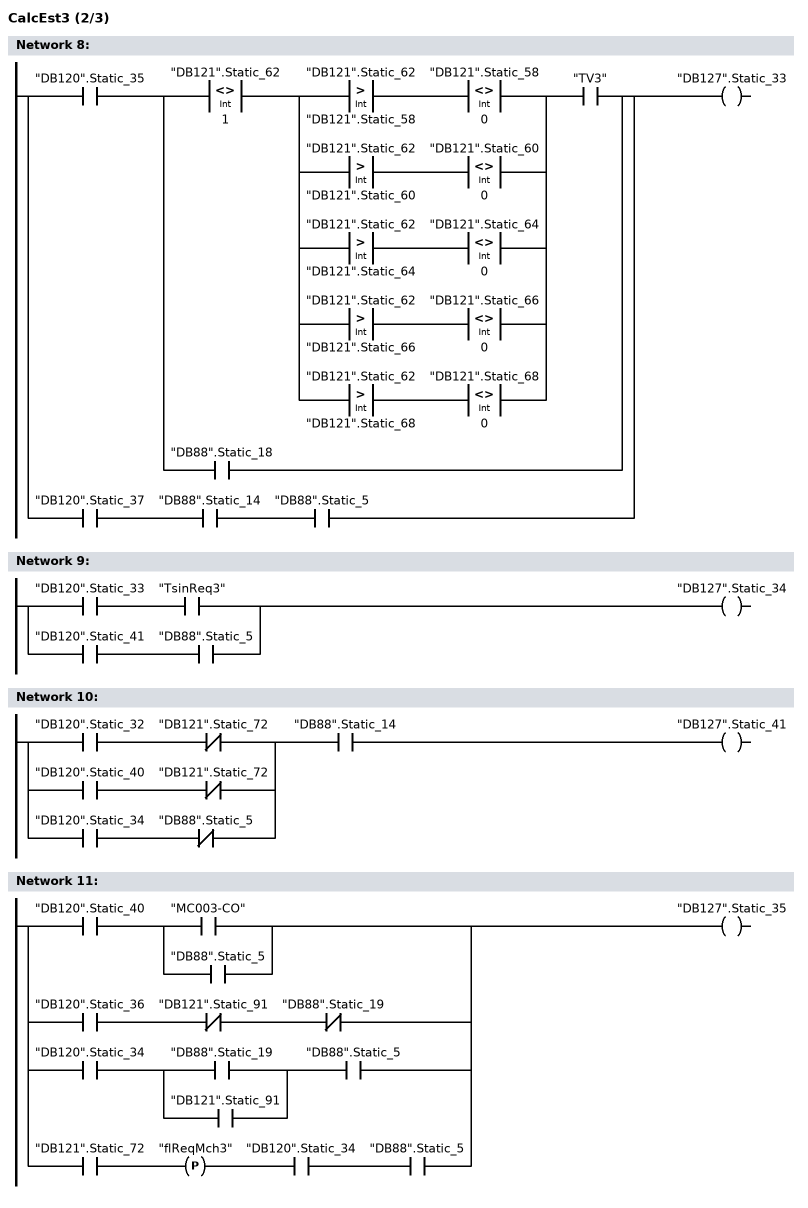
   "DB127".Static_33 := ("DB120".Static_35 AND ((("DB121".Static_62 <> 1) AND ((("DB121".Static_62 > "DB121".Static_58) AND ("DB121".Static_58 <> 0)) OR (("DB121".Static_62 > "DB121".Static_60) AND ("DB121".Static_60 <> 0)) OR (("DB121".Static_62 > "DB121".Static_64) AND ("DB121".Static_64 <> 0)) OR (("DB121".Static_62 > "DB121".Static_66) AND ("DB121".Static_66 <> 0)) OR (("DB121".Static_62 > "DB121".Static_68) AND ("DB121".Static_68 <> 0))) AND "TV3") OR "DB88".Static_18)) OR ("DB120".Static_37 AND "DB88".Static_14 AND "DB88".Static_5);
END_REGION

REGION Network 9
   RUNG wire#powerrail
      Contact( "DB120".Static_33 )
      Contact( "TsinReq3" )
      wire#w1
      Coil( "DB127".Static_34 )
   END_RUNG
   RUNG wire#powerrail
      Contact( "DB120".Static_41 )
      Contact( "DB88".Static_5 )
   END_RUNG wire#w1
   // the same network as SCL:
   "DB127".Static_34 := ("DB120".Static_33 AND "TsinReq3") OR ("DB120".Static_41 AND "DB88".Static_5);
END_REGION

REGION Network 10
   RUNG wire#powerrail
      Contact( "DB120".Static_32 )
      I_Contact( "DB121".Static_72 )
      wire#w1
      Contact( "DB88".Static_14 )
      Coil( "DB127".Static_41 )
   END_RUNG
   RUNG wire#powerrail
      Contact( "DB120".Static_40 )
      I_Contact( "DB121".Static_72 )
   END_RUNG wire#w1
   RUNG wire#powerrail
      Contact( "DB120".Static_34 )
      I_Contact( "DB88".Static_5 )
   END_RUNG wire#w1
   // the same network as SCL:
   "DB127".Static_41 := (("DB120".Static_32 AND NOT "DB121".Static_72) OR ("DB120".Static_40 AND NOT "DB121".Static_72) OR ("DB120".Static_34 AND NOT "DB88".Static_5)) AND "DB88".Static_14;
END_REGION

REGION Network 11
   #_w1 := "DB121".Static_72 AND NOT "flReqMch3";   // rising edge
   "flReqMch3" := "DB121".Static_72;
   "DB127".Static_35 := ("DB120".Static_40 AND ("MC003-CO" OR "DB88".Static_5)) OR ("DB120".Static_36 AND NOT "DB121".Static_91 AND NOT "DB88".Static_19) OR ("DB120".Static_34 AND ("DB88".Static_19 OR "DB121".Static_91) AND "DB88".Static_5) OR (#_w1 AND "DB120".Static_34 AND "DB88".Static_5);
END_REGION

REGION Network 12
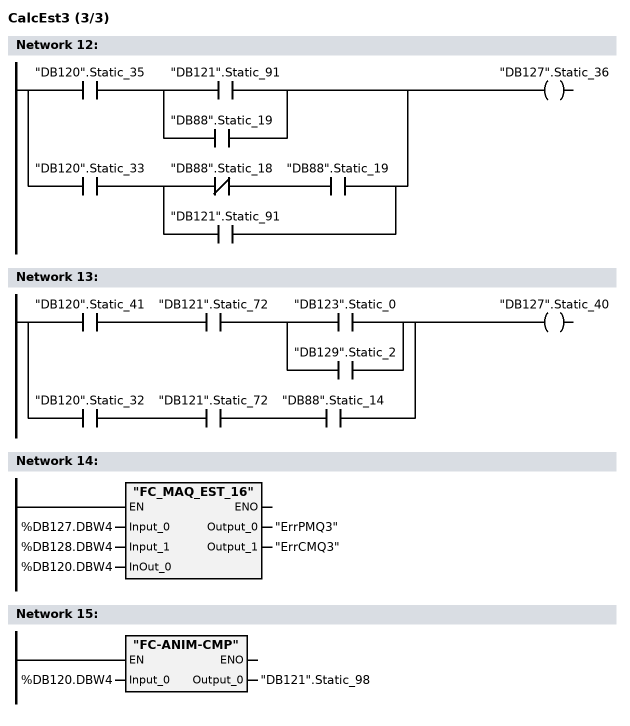
   "DB127".Static_36 := ("DB120".Static_35 AND ("DB121".Static_91 OR "DB88".Static_19)) OR ("DB120".Static_33 AND ("DB121".Static_91 OR (NOT "DB88".Static_18 AND "DB88".Static_19)));
END_REGION

REGION Network 13
   "DB127".Static_40 := ("DB120".Static_41 AND "DB121".Static_72 AND ("DB123".Static_0 OR "DB129".Static_2)) OR ("DB120".Static_32 AND "DB121".Static_72 AND "DB88".Static_14);
END_REGION

REGION Network 14
   RUNG wire#powerrail
      "FC_MAQ_EST_16"(Input_0 := %DB127.DBW4, Input_1 := %DB128.DBW4, Output_0 => "ErrPMQ3", Output_1 => "ErrCMQ3", InOut_0 := %DB120.DBW4)
   END_RUNG
   // the same network as SCL:
   "FC_MAQ_EST_16"(Input_0 := %DB127.DBW4,
                   Input_1 := %DB128.DBW4,
                   InOut_0 := %DB120.DBW4,
                   Output_0 => "ErrPMQ3",
                   Output_1 => "ErrCMQ3");
END_REGION

REGION Network 15
   RUNG wire#powerrail
      "FC-ANIM-CMP"(Input_0 := %DB120.DBW4, Output_0 => "DB121".Static_98)
   END_RUNG
   // the same network as SCL:
   "FC-ANIM-CMP"(Input_0 := %DB120.DBW4, Output_0 => "DB121".Static_98);
END_REGION
END_FUNCTION

FUNCTION "CalcEst4" : Void   // FC39, LAD
{ S7_Optimized_Access := 'FALSE' }
VERSION : 0.1
   VAR_TEMP   // added for the SCL form of the ladder/FBD networks
      _w1 : Bool;
   END_VAR
BEGIN

REGION Network 1
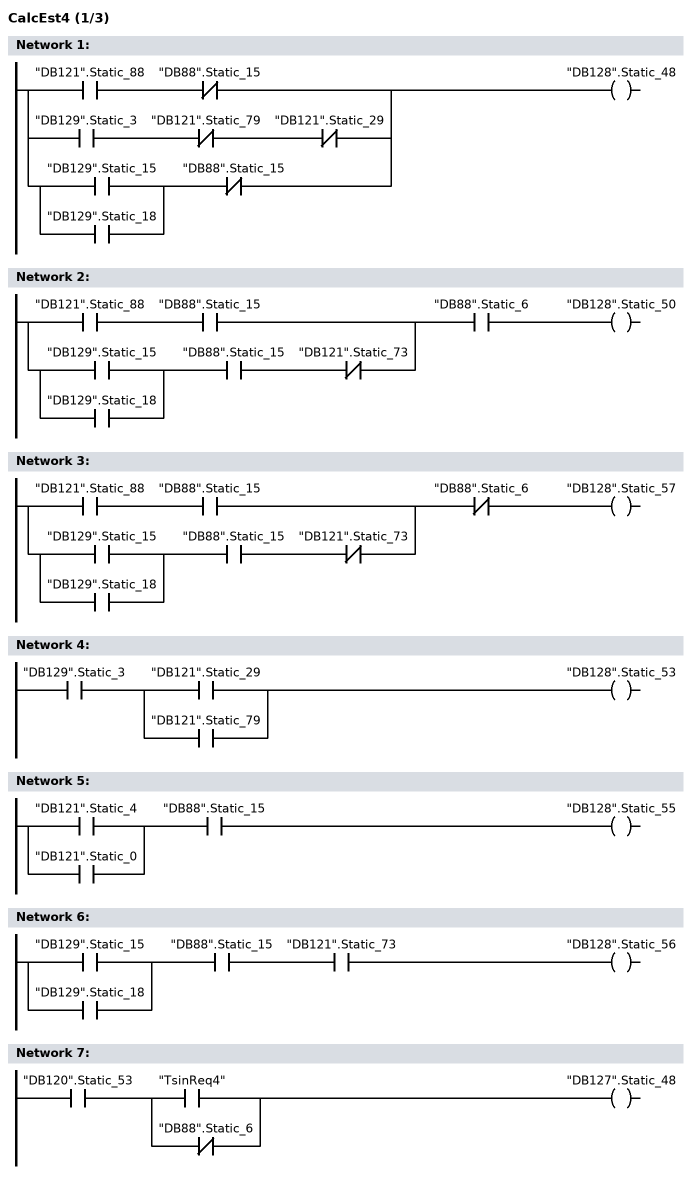
   RUNG wire#powerrail
      Contact( "DB121".Static_88 )
      I_Contact( "DB88".Static_15 )
      wire#w1
      Coil( "DB128".Static_48 )
   END_RUNG
   RUNG wire#powerrail
      Contact( "DB129".Static_3 )
      I_Contact( "DB121".Static_79 )
      I_Contact( "DB121".Static_29 )
   END_RUNG wire#w1
   RUNG wire#powerrail
      Contact( "DB129".Static_15 )
      wire#w2
      I_Contact( "DB88".Static_15 )
   END_RUNG wire#w1
   RUNG wire#powerrail
      Contact( "DB129".Static_18 )
   END_RUNG wire#w2
   // the same network as SCL:
   "DB128".Static_48 := ("DB121".Static_88 AND NOT "DB88".Static_15) OR ("DB129".Static_3 AND NOT "DB121".Static_79 AND NOT "DB121".Static_29) OR (("DB129".Static_15 OR "DB129".Static_18) AND NOT "DB88".Static_15);
END_REGION

REGION Network 2
   RUNG wire#powerrail
      Contact( "DB121".Static_88 )
      Contact( "DB88".Static_15 )
      wire#w1
      Contact( "DB88".Static_6 )
      Coil( "DB128".Static_50 )
   END_RUNG
   RUNG wire#powerrail
      Contact( "DB129".Static_15 )
      wire#w2
      Contact( "DB88".Static_15 )
      I_Contact( "DB121".Static_73 )
   END_RUNG wire#w1
   RUNG wire#powerrail
      Contact( "DB129".Static_18 )
   END_RUNG wire#w2
   // the same network as SCL:
   "DB128".Static_50 := (("DB121".Static_88 AND "DB88".Static_15) OR (("DB129".Static_15 OR "DB129".Static_18) AND "DB88".Static_15 AND NOT "DB121".Static_73)) AND "DB88".Static_6;
END_REGION

REGION Network 3
   RUNG wire#powerrail
      Contact( "DB121".Static_88 )
      Contact( "DB88".Static_15 )
      wire#w1
      I_Contact( "DB88".Static_6 )
      Coil( "DB128".Static_57 )
   END_RUNG
   RUNG wire#powerrail
      Contact( "DB129".Static_15 )
      wire#w2
      Contact( "DB88".Static_15 )
      I_Contact( "DB121".Static_73 )
   END_RUNG wire#w1
   RUNG wire#powerrail
      Contact( "DB129".Static_18 )
   END_RUNG wire#w2
   // the same network as SCL:
   "DB128".Static_57 := (("DB121".Static_88 AND "DB88".Static_15) OR (("DB129".Static_15 OR "DB129".Static_18) AND "DB88".Static_15 AND NOT "DB121".Static_73)) AND NOT "DB88".Static_6;
END_REGION

REGION Network 4
   "DB128".Static_53 := "DB129".Static_3 AND ("DB121".Static_29 OR "DB121".Static_79);
END_REGION

REGION Network 5
   RUNG wire#powerrail
      Contact( "DB121".Static_4 )
      wire#w1
      Contact( "DB88".Static_15 )
      Coil( "DB128".Static_55 )
   END_RUNG
   RUNG wire#powerrail
      Contact( "DB121".Static_0 )
   END_RUNG wire#w1
   // the same network as SCL:
   "DB128".Static_55 := ("DB121".Static_4 OR "DB121".Static_0) AND "DB88".Static_15;
END_REGION

REGION Network 6
   RUNG wire#powerrail
      Contact( "DB129".Static_15 )
      wire#w1
      Contact( "DB88".Static_15 )
      Contact( "DB121".Static_73 )
      Coil( "DB128".Static_56 )
   END_RUNG
   RUNG wire#powerrail
      Contact( "DB129".Static_18 )
   END_RUNG wire#w1
   // the same network as SCL:
   "DB128".Static_56 := ("DB129".Static_15 OR "DB129".Static_18) AND "DB88".Static_15 AND "DB121".Static_73;
END_REGION

REGION Network 7
   "DB127".Static_48 := "DB120".Static_53 AND ("TsinReq4" OR NOT "DB88".Static_6);
END_REGION

REGION Network 8
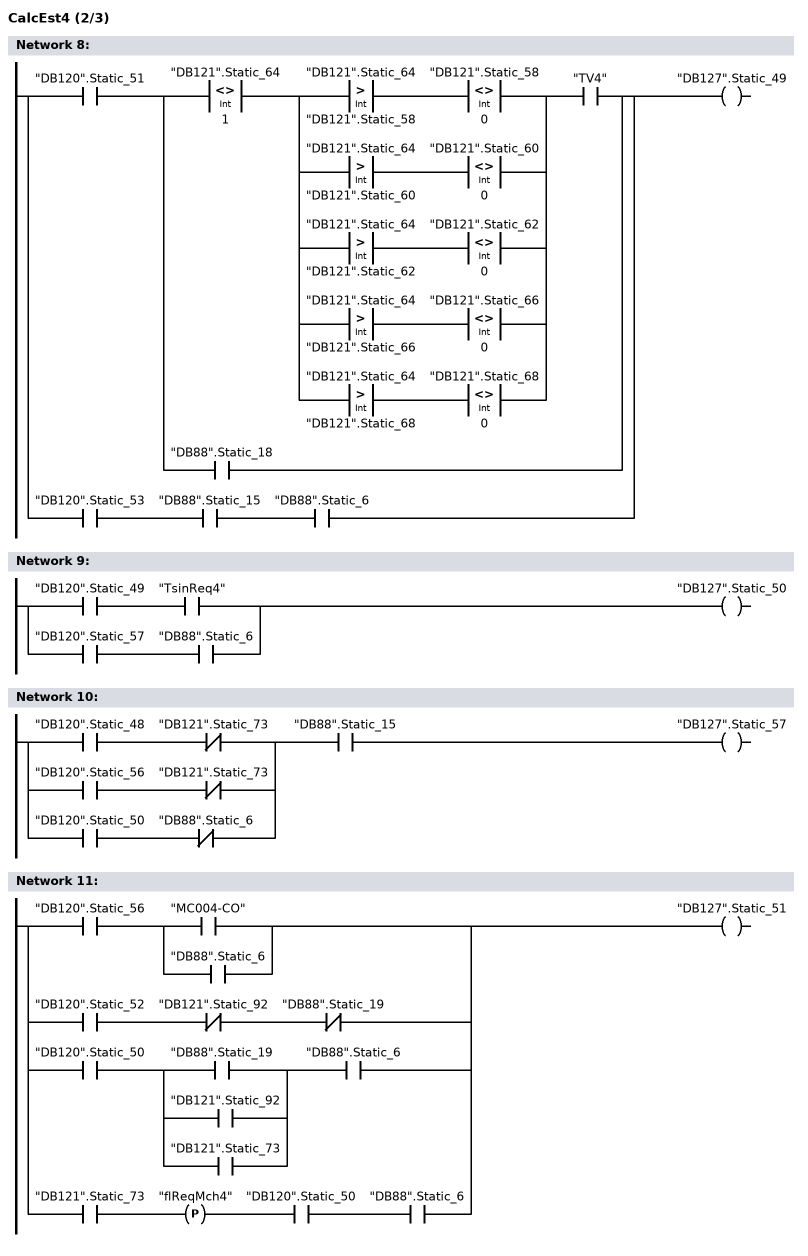
   "DB127".Static_49 := ("DB120".Static_51 AND ((("DB121".Static_64 <> 1) AND ((("DB121".Static_64 > "DB121".Static_58) AND ("DB121".Static_58 <> 0)) OR (("DB121".Static_64 > "DB121".Static_60) AND ("DB121".Static_60 <> 0)) OR (("DB121".Static_64 > "DB121".Static_62) AND ("DB121".Static_62 <> 0)) OR (("DB121".Static_64 > "DB121".Static_66) AND ("DB121".Static_66 <> 0)) OR (("DB121".Static_64 > "DB121".Static_68) AND ("DB121".Static_68 <> 0))) AND "TV4") OR "DB88".Static_18)) OR ("DB120".Static_53 AND "DB88".Static_15 AND "DB88".Static_6);
END_REGION

REGION Network 9
   RUNG wire#powerrail
      Contact( "DB120".Static_49 )
      Contact( "TsinReq4" )
      wire#w1
      Coil( "DB127".Static_50 )
   END_RUNG
   RUNG wire#powerrail
      Contact( "DB120".Static_57 )
      Contact( "DB88".Static_6 )
   END_RUNG wire#w1
   // the same network as SCL:
   "DB127".Static_50 := ("DB120".Static_49 AND "TsinReq4") OR ("DB120".Static_57 AND "DB88".Static_6);
END_REGION

REGION Network 10
   RUNG wire#powerrail
      Contact( "DB120".Static_48 )
      I_Contact( "DB121".Static_73 )
      wire#w1
      Contact( "DB88".Static_15 )
      Coil( "DB127".Static_57 )
   END_RUNG
   RUNG wire#powerrail
      Contact( "DB120".Static_56 )
      I_Contact( "DB121".Static_73 )
   END_RUNG wire#w1
   RUNG wire#powerrail
      Contact( "DB120".Static_50 )
      I_Contact( "DB88".Static_6 )
   END_RUNG wire#w1
   // the same network as SCL:
   "DB127".Static_57 := (("DB120".Static_48 AND NOT "DB121".Static_73) OR ("DB120".Static_56 AND NOT "DB121".Static_73) OR ("DB120".Static_50 AND NOT "DB88".Static_6)) AND "DB88".Static_15;
END_REGION

REGION Network 11
   #_w1 := "DB121".Static_73 AND NOT "flReqMch4";   // rising edge
   "flReqMch4" := "DB121".Static_73;
   "DB127".Static_51 := ("DB120".Static_56 AND ("MC004-CO" OR "DB88".Static_6)) OR ("DB120".Static_52 AND NOT "DB121".Static_92 AND NOT "DB88".Static_19) OR ("DB120".Static_50 AND ("DB88".Static_19 OR "DB121".Static_92 OR "DB121".Static_73) AND "DB88".Static_6) OR (#_w1 AND "DB120".Static_50 AND "DB88".Static_6);
END_REGION

REGION Network 12
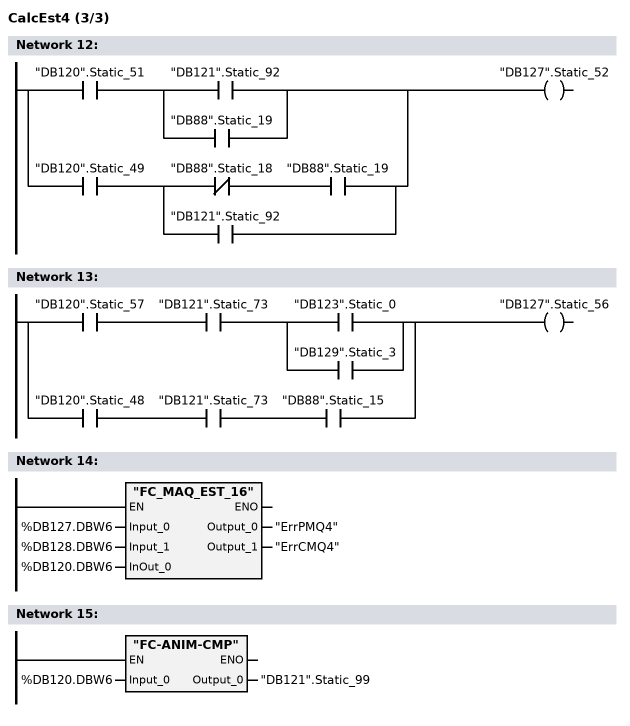
   "DB127".Static_52 := ("DB120".Static_51 AND ("DB121".Static_92 OR "DB88".Static_19)) OR ("DB120".Static_49 AND ("DB121".Static_92 OR (NOT "DB88".Static_18 AND "DB88".Static_19)));
END_REGION

REGION Network 13
   "DB127".Static_56 := ("DB120".Static_57 AND "DB121".Static_73 AND ("DB123".Static_0 OR "DB129".Static_3)) OR ("DB120".Static_48 AND "DB121".Static_73 AND "DB88".Static_15);
END_REGION

REGION Network 14
   RUNG wire#powerrail
      "FC_MAQ_EST_16"(Input_0 := %DB127.DBW6, Input_1 := %DB128.DBW6, Output_0 => "ErrPMQ4", Output_1 => "ErrCMQ4", InOut_0 := %DB120.DBW6)
   END_RUNG
   // the same network as SCL:
   "FC_MAQ_EST_16"(Input_0 := %DB127.DBW6,
                   Input_1 := %DB128.DBW6,
                   InOut_0 := %DB120.DBW6,
                   Output_0 => "ErrPMQ4",
                   Output_1 => "ErrCMQ4");
END_REGION

REGION Network 15
   RUNG wire#powerrail
      "FC-ANIM-CMP"(Input_0 := %DB120.DBW6, Output_0 => "DB121".Static_99)
   END_RUNG
   // the same network as SCL:
   "FC-ANIM-CMP"(Input_0 := %DB120.DBW6, Output_0 => "DB121".Static_99);
END_REGION
END_FUNCTION

FUNCTION "CalcEst5" : Void   // FC40, LAD
{ S7_Optimized_Access := 'FALSE' }
VERSION : 0.1
   VAR_TEMP   // added for the SCL form of the ladder/FBD networks
      _w1 : Bool;
   END_VAR
BEGIN

REGION Network 1
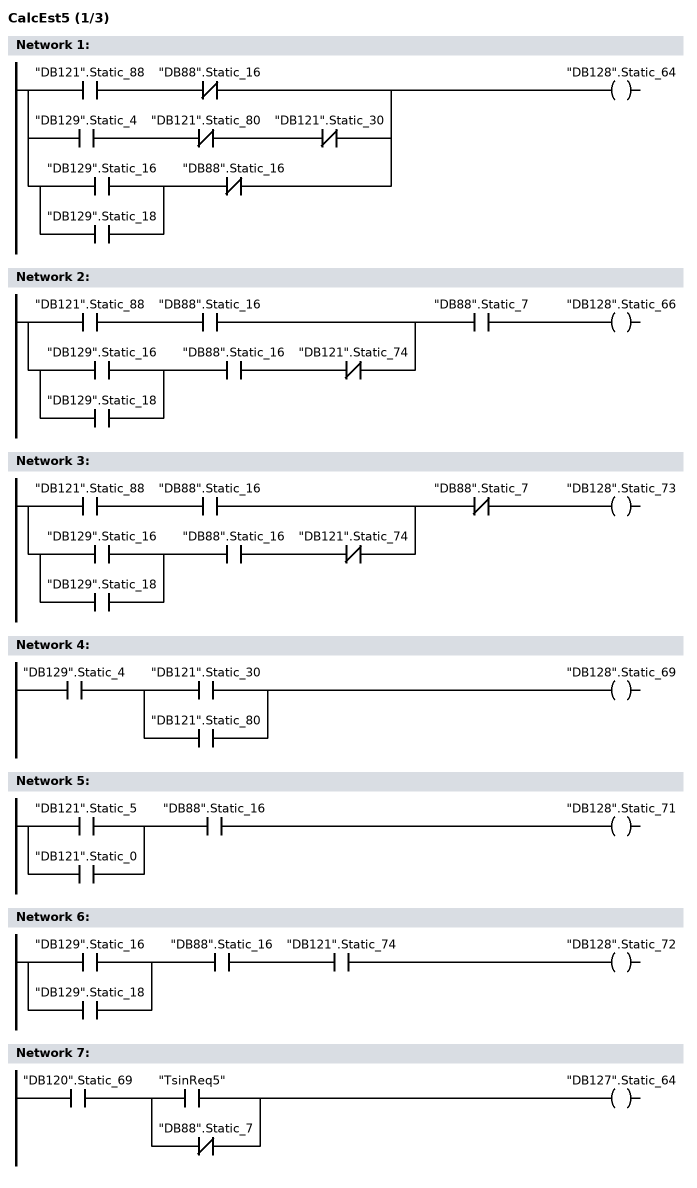
   RUNG wire#powerrail
      Contact( "DB121".Static_88 )
      I_Contact( "DB88".Static_16 )
      wire#w1
      Coil( "DB128".Static_64 )
   END_RUNG
   RUNG wire#powerrail
      Contact( "DB129".Static_4 )
      I_Contact( "DB121".Static_80 )
      I_Contact( "DB121".Static_30 )
   END_RUNG wire#w1
   RUNG wire#powerrail
      Contact( "DB129".Static_16 )
      wire#w2
      I_Contact( "DB88".Static_16 )
   END_RUNG wire#w1
   RUNG wire#powerrail
      Contact( "DB129".Static_18 )
   END_RUNG wire#w2
   // the same network as SCL:
   "DB128".Static_64 := ("DB121".Static_88 AND NOT "DB88".Static_16) OR ("DB129".Static_4 AND NOT "DB121".Static_80 AND NOT "DB121".Static_30) OR (("DB129".Static_16 OR "DB129".Static_18) AND NOT "DB88".Static_16);
END_REGION

REGION Network 2
   RUNG wire#powerrail
      Contact( "DB121".Static_88 )
      Contact( "DB88".Static_16 )
      wire#w1
      Contact( "DB88".Static_7 )
      Coil( "DB128".Static_66 )
   END_RUNG
   RUNG wire#powerrail
      Contact( "DB129".Static_16 )
      wire#w2
      Contact( "DB88".Static_16 )
      I_Contact( "DB121".Static_74 )
   END_RUNG wire#w1
   RUNG wire#powerrail
      Contact( "DB129".Static_18 )
   END_RUNG wire#w2
   // the same network as SCL:
   "DB128".Static_66 := (("DB121".Static_88 AND "DB88".Static_16) OR (("DB129".Static_16 OR "DB129".Static_18) AND "DB88".Static_16 AND NOT "DB121".Static_74)) AND "DB88".Static_7;
END_REGION

REGION Network 3
   RUNG wire#powerrail
      Contact( "DB121".Static_88 )
      Contact( "DB88".Static_16 )
      wire#w1
      I_Contact( "DB88".Static_7 )
      Coil( "DB128".Static_73 )
   END_RUNG
   RUNG wire#powerrail
      Contact( "DB129".Static_16 )
      wire#w2
      Contact( "DB88".Static_16 )
      I_Contact( "DB121".Static_74 )
   END_RUNG wire#w1
   RUNG wire#powerrail
      Contact( "DB129".Static_18 )
   END_RUNG wire#w2
   // the same network as SCL:
   "DB128".Static_73 := (("DB121".Static_88 AND "DB88".Static_16) OR (("DB129".Static_16 OR "DB129".Static_18) AND "DB88".Static_16 AND NOT "DB121".Static_74)) AND NOT "DB88".Static_7;
END_REGION

REGION Network 4
   "DB128".Static_69 := "DB129".Static_4 AND ("DB121".Static_30 OR "DB121".Static_80);
END_REGION

REGION Network 5
   RUNG wire#powerrail
      Contact( "DB121".Static_5 )
      wire#w1
      Contact( "DB88".Static_16 )
      Coil( "DB128".Static_71 )
   END_RUNG
   RUNG wire#powerrail
      Contact( "DB121".Static_0 )
   END_RUNG wire#w1
   // the same network as SCL:
   "DB128".Static_71 := ("DB121".Static_5 OR "DB121".Static_0) AND "DB88".Static_16;
END_REGION

REGION Network 6
   RUNG wire#powerrail
      Contact( "DB129".Static_16 )
      wire#w1
      Contact( "DB88".Static_16 )
      Contact( "DB121".Static_74 )
      Coil( "DB128".Static_72 )
   END_RUNG
   RUNG wire#powerrail
      Contact( "DB129".Static_18 )
   END_RUNG wire#w1
   // the same network as SCL:
   "DB128".Static_72 := ("DB129".Static_16 OR "DB129".Static_18) AND "DB88".Static_16 AND "DB121".Static_74;
END_REGION

REGION Network 7
   "DB127".Static_64 := "DB120".Static_69 AND ("TsinReq5" OR NOT "DB88".Static_7);
END_REGION

REGION Network 8
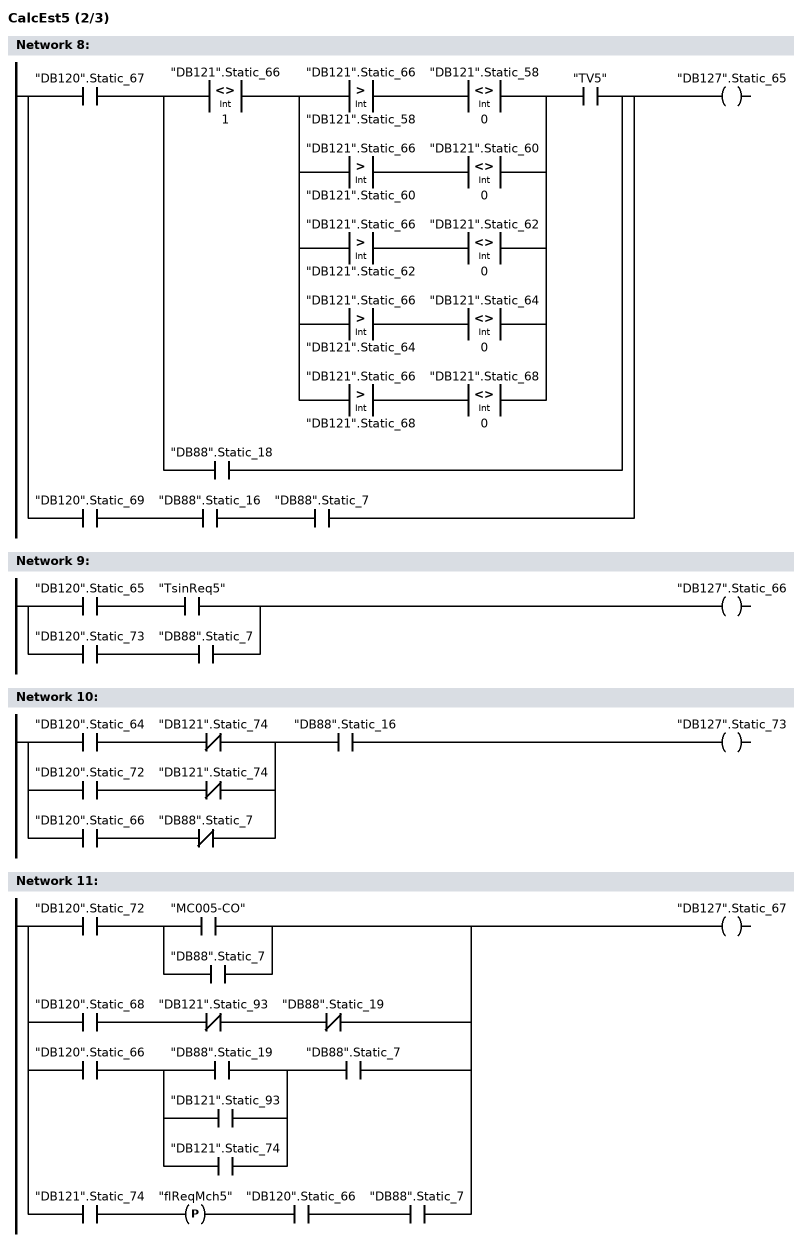
   "DB127".Static_65 := ("DB120".Static_67 AND ((("DB121".Static_66 <> 1) AND ((("DB121".Static_66 > "DB121".Static_58) AND ("DB121".Static_58 <> 0)) OR (("DB121".Static_66 > "DB121".Static_60) AND ("DB121".Static_60 <> 0)) OR (("DB121".Static_66 > "DB121".Static_62) AND ("DB121".Static_62 <> 0)) OR (("DB121".Static_66 > "DB121".Static_64) AND ("DB121".Static_64 <> 0)) OR (("DB121".Static_66 > "DB121".Static_68) AND ("DB121".Static_68 <> 0))) AND "TV5") OR "DB88".Static_18)) OR ("DB120".Static_69 AND "DB88".Static_16 AND "DB88".Static_7);
END_REGION

REGION Network 9
   RUNG wire#powerrail
      Contact( "DB120".Static_65 )
      Contact( "TsinReq5" )
      wire#w1
      Coil( "DB127".Static_66 )
   END_RUNG
   RUNG wire#powerrail
      Contact( "DB120".Static_73 )
      Contact( "DB88".Static_7 )
   END_RUNG wire#w1
   // the same network as SCL:
   "DB127".Static_66 := ("DB120".Static_65 AND "TsinReq5") OR ("DB120".Static_73 AND "DB88".Static_7);
END_REGION

REGION Network 10
   RUNG wire#powerrail
      Contact( "DB120".Static_64 )
      I_Contact( "DB121".Static_74 )
      wire#w1
      Contact( "DB88".Static_16 )
      Coil( "DB127".Static_73 )
   END_RUNG
   RUNG wire#powerrail
      Contact( "DB120".Static_72 )
      I_Contact( "DB121".Static_74 )
   END_RUNG wire#w1
   RUNG wire#powerrail
      Contact( "DB120".Static_66 )
      I_Contact( "DB88".Static_7 )
   END_RUNG wire#w1
   // the same network as SCL:
   "DB127".Static_73 := (("DB120".Static_64 AND NOT "DB121".Static_74) OR ("DB120".Static_72 AND NOT "DB121".Static_74) OR ("DB120".Static_66 AND NOT "DB88".Static_7)) AND "DB88".Static_16;
END_REGION

REGION Network 11
   #_w1 := "DB121".Static_74 AND NOT "flReqMch5";   // rising edge
   "flReqMch5" := "DB121".Static_74;
   "DB127".Static_67 := ("DB120".Static_72 AND ("MC005-CO" OR "DB88".Static_7)) OR ("DB120".Static_68 AND NOT "DB121".Static_93 AND NOT "DB88".Static_19) OR ("DB120".Static_66 AND ("DB88".Static_19 OR "DB121".Static_93 OR "DB121".Static_74) AND "DB88".Static_7) OR (#_w1 AND "DB120".Static_66 AND "DB88".Static_7);
END_REGION

REGION Network 12
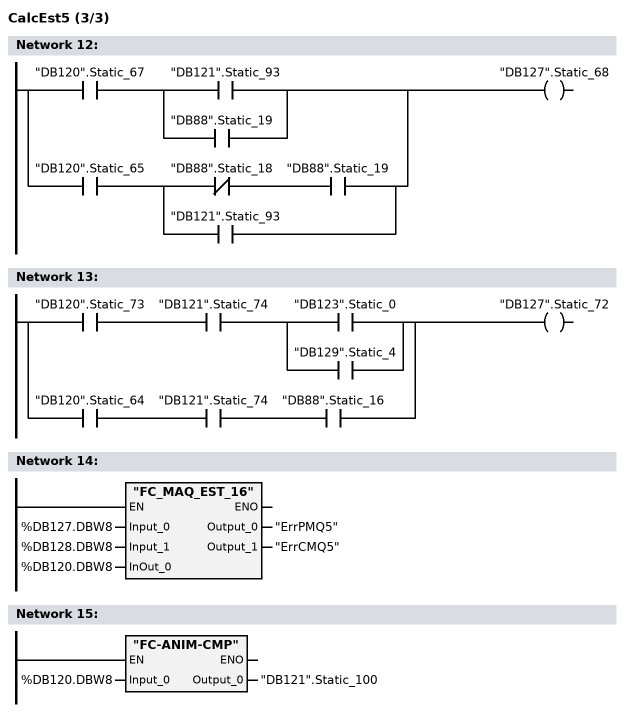
   "DB127".Static_68 := ("DB120".Static_67 AND ("DB121".Static_93 OR "DB88".Static_19)) OR ("DB120".Static_65 AND ("DB121".Static_93 OR (NOT "DB88".Static_18 AND "DB88".Static_19)));
END_REGION

REGION Network 13
   "DB127".Static_72 := ("DB120".Static_73 AND "DB121".Static_74 AND ("DB123".Static_0 OR "DB129".Static_4)) OR ("DB120".Static_64 AND "DB121".Static_74 AND "DB88".Static_16);
END_REGION

REGION Network 14
   RUNG wire#powerrail
      "FC_MAQ_EST_16"(Input_0 := %DB127.DBW8, Input_1 := %DB128.DBW8, Output_0 => "ErrPMQ5", Output_1 => "ErrCMQ5", InOut_0 := %DB120.DBW8)
   END_RUNG
   // the same network as SCL:
   "FC_MAQ_EST_16"(Input_0 := %DB127.DBW8,
                   Input_1 := %DB128.DBW8,
                   InOut_0 := %DB120.DBW8,
                   Output_0 => "ErrPMQ5",
                   Output_1 => "ErrCMQ5");
END_REGION

REGION Network 15
   RUNG wire#powerrail
      "FC-ANIM-CMP"(Input_0 := %DB120.DBW8, Output_0 => "DB121".Static_100)
   END_RUNG
   // the same network as SCL:
   "FC-ANIM-CMP"(Input_0 := %DB120.DBW8, Output_0 => "DB121".Static_100);
END_REGION
END_FUNCTION

FUNCTION "CalcEst0" : Void   // FC42, LAD
{ S7_Optimized_Access := 'FALSE' }
VERSION : 0.1
BEGIN

REGION Network 1
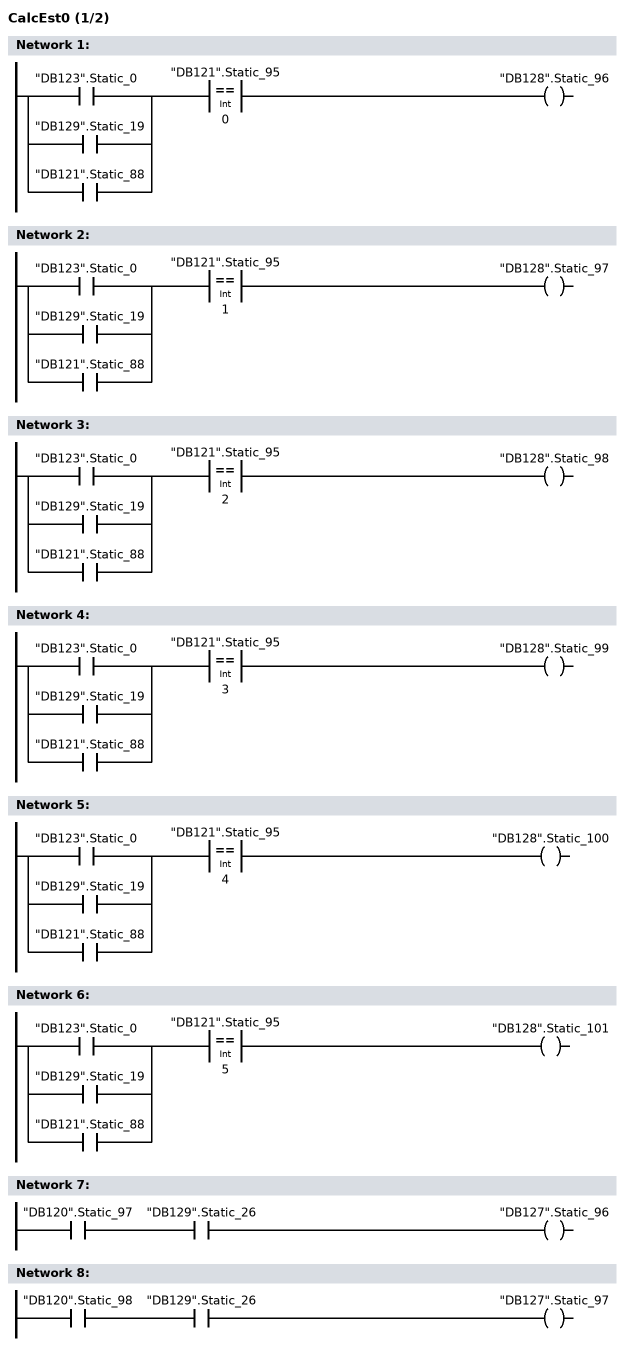
   RUNG wire#powerrail
      Contact( "DB123".Static_0 )
      wire#w1
      { S7_Templates := "SrcType := Int" } EQ_Contact(in1 := "DB121".Static_95, in2 := 0)
      Coil( "DB128".Static_96 )
   END_RUNG
   RUNG wire#powerrail
      Contact( "DB129".Static_19 )
   END_RUNG wire#w1
   RUNG wire#powerrail
      Contact( "DB121".Static_88 )
   END_RUNG wire#w1
   // the same network as SCL:
   "DB128".Static_96 := ("DB123".Static_0 OR "DB129".Static_19 OR "DB121".Static_88) AND ("DB121".Static_95 = 0);
END_REGION

REGION Network 2
   RUNG wire#powerrail
      Contact( "DB123".Static_0 )
      wire#w1
      { S7_Templates := "SrcType := Int" } EQ_Contact(in1 := "DB121".Static_95, in2 := 1)
      Coil( "DB128".Static_97 )
   END_RUNG
   RUNG wire#powerrail
      Contact( "DB129".Static_19 )
   END_RUNG wire#w1
   RUNG wire#powerrail
      Contact( "DB121".Static_88 )
   END_RUNG wire#w1
   // the same network as SCL:
   "DB128".Static_97 := ("DB123".Static_0 OR "DB129".Static_19 OR "DB121".Static_88) AND ("DB121".Static_95 = 1);
END_REGION

REGION Network 3
   RUNG wire#powerrail
      Contact( "DB123".Static_0 )
      wire#w1
      { S7_Templates := "SrcType := Int" } EQ_Contact(in1 := "DB121".Static_95, in2 := 2)
      Coil( "DB128".Static_98 )
   END_RUNG
   RUNG wire#powerrail
      Contact( "DB129".Static_19 )
   END_RUNG wire#w1
   RUNG wire#powerrail
      Contact( "DB121".Static_88 )
   END_RUNG wire#w1
   // the same network as SCL:
   "DB128".Static_98 := ("DB123".Static_0 OR "DB129".Static_19 OR "DB121".Static_88) AND ("DB121".Static_95 = 2);
END_REGION

REGION Network 4
   RUNG wire#powerrail
      Contact( "DB123".Static_0 )
      wire#w1
      { S7_Templates := "SrcType := Int" } EQ_Contact(in1 := "DB121".Static_95, in2 := 3)
      Coil( "DB128".Static_99 )
   END_RUNG
   RUNG wire#powerrail
      Contact( "DB129".Static_19 )
   END_RUNG wire#w1
   RUNG wire#powerrail
      Contact( "DB121".Static_88 )
   END_RUNG wire#w1
   // the same network as SCL:
   "DB128".Static_99 := ("DB123".Static_0 OR "DB129".Static_19 OR "DB121".Static_88) AND ("DB121".Static_95 = 3);
END_REGION

REGION Network 5
   RUNG wire#powerrail
      Contact( "DB123".Static_0 )
      wire#w1
      { S7_Templates := "SrcType := Int" } EQ_Contact(in1 := "DB121".Static_95, in2 := 4)
      Coil( "DB128".Static_100 )
   END_RUNG
   RUNG wire#powerrail
      Contact( "DB129".Static_19 )
   END_RUNG wire#w1
   RUNG wire#powerrail
      Contact( "DB121".Static_88 )
   END_RUNG wire#w1
   // the same network as SCL:
   "DB128".Static_100 := ("DB123".Static_0 OR "DB129".Static_19 OR "DB121".Static_88) AND ("DB121".Static_95 = 4);
END_REGION

REGION Network 6
   RUNG wire#powerrail
      Contact( "DB123".Static_0 )
      wire#w1
      { S7_Templates := "SrcType := Int" } EQ_Contact(in1 := "DB121".Static_95, in2 := 5)
      Coil( "DB128".Static_101 )
   END_RUNG
   RUNG wire#powerrail
      Contact( "DB129".Static_19 )
   END_RUNG wire#w1
   RUNG wire#powerrail
      Contact( "DB121".Static_88 )
   END_RUNG wire#w1
   // the same network as SCL:
   "DB128".Static_101 := ("DB123".Static_0 OR "DB129".Static_19 OR "DB121".Static_88) AND ("DB121".Static_95 = 5);
END_REGION

REGION Network 7
   RUNG wire#powerrail
      Contact( "DB120".Static_97 )
      Contact( "DB129".Static_26 )
      Coil( "DB127".Static_96 )
   END_RUNG
   // the same network as SCL:
   "DB127".Static_96 := "DB120".Static_97 AND "DB129".Static_26;
END_REGION

REGION Network 8
   RUNG wire#powerrail
      Contact( "DB120".Static_98 )
      Contact( "DB129".Static_26 )
      Coil( "DB127".Static_97 )
   END_RUNG
   // the same network as SCL:
   "DB127".Static_97 := "DB120".Static_98 AND "DB129".Static_26;
END_REGION

REGION Network 9
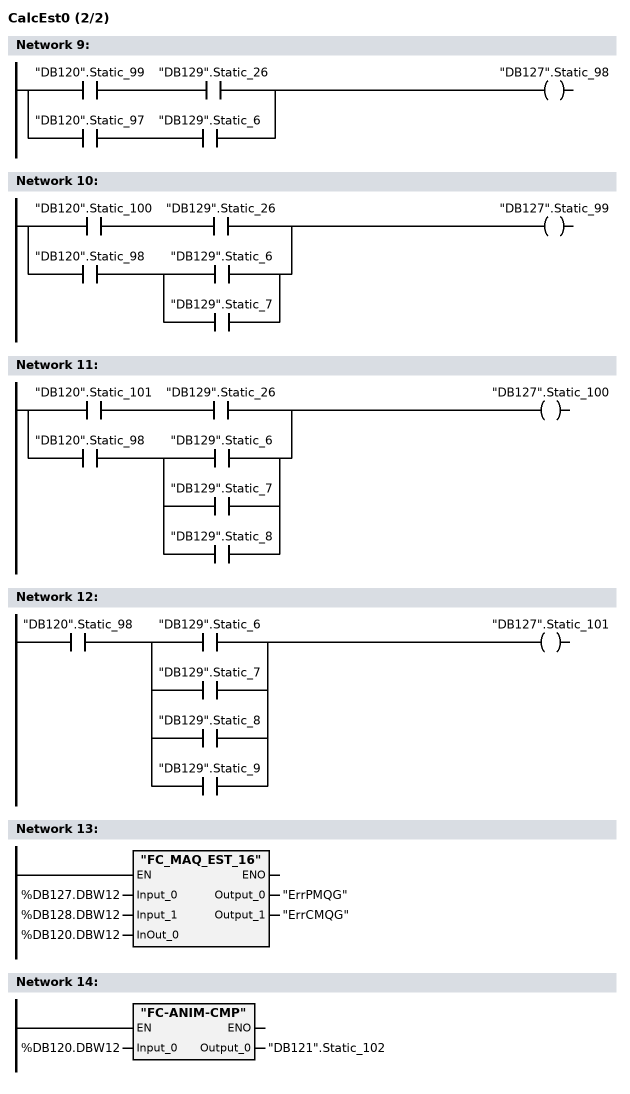
   RUNG wire#powerrail
      Contact( "DB120".Static_99 )
      Contact( "DB129".Static_26 )
      wire#w1
      Coil( "DB127".Static_98 )
   END_RUNG
   RUNG wire#powerrail
      Contact( "DB120".Static_97 )
      Contact( "DB129".Static_6 )
   END_RUNG wire#w1
   // the same network as SCL:
   "DB127".Static_98 := ("DB120".Static_99 AND "DB129".Static_26) OR ("DB120".Static_97 AND "DB129".Static_6);
END_REGION

REGION Network 10
   "DB127".Static_99 := ("DB120".Static_100 AND "DB129".Static_26) OR ("DB120".Static_98 AND ("DB129".Static_6 OR "DB129".Static_7));
END_REGION

REGION Network 11
   "DB127".Static_100 := ("DB120".Static_101 AND "DB129".Static_26) OR ("DB120".Static_98 AND ("DB129".Static_6 OR "DB129".Static_7 OR "DB129".Static_8));
END_REGION

REGION Network 12
   "DB127".Static_101 := "DB120".Static_98 AND ("DB129".Static_6 OR "DB129".Static_7 OR "DB129".Static_8 OR "DB129".Static_9);
END_REGION

REGION Network 13
   RUNG wire#powerrail
      "FC_MAQ_EST_16"(Input_0 := %DB127.DBW12, Input_1 := %DB128.DBW12, Output_0 => "ErrPMQG", Output_1 => "ErrCMQG", InOut_0 := %DB120.DBW12)
   END_RUNG
   // the same network as SCL:
   "FC_MAQ_EST_16"(Input_0 := %DB127.DBW12,
                   Input_1 := %DB128.DBW12,
                   InOut_0 := %DB120.DBW12,
                   Output_0 => "ErrPMQG",
                   Output_1 => "ErrCMQG");
END_REGION

REGION Network 14
   RUNG wire#powerrail
      "FC-ANIM-CMP"(Input_0 := %DB120.DBW12, Output_0 => "DB121".Static_102)
   END_RUNG
   // the same network as SCL:
   "FC-ANIM-CMP"(Input_0 := %DB120.DBW12, Output_0 => "DB121".Static_102);
END_REGION
END_FUNCTION

FUNCTION "CorreccReqCmpAlta" : Void   // FC44, LAD
{ S7_Optimized_Access := 'FALSE' }
VERSION : 0.1
BEGIN

REGION Network 1
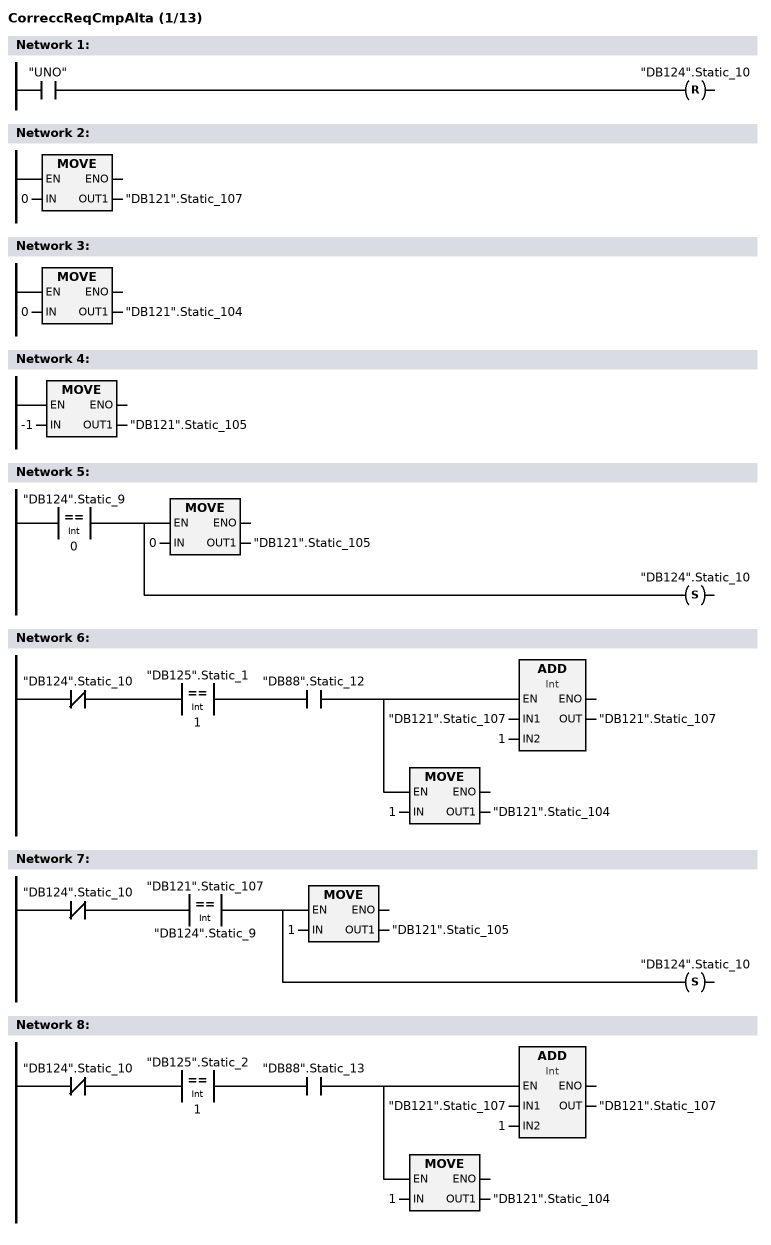
   RUNG wire#powerrail
      Contact( "UNO" )
      R_Coil( "DB124".Static_10 )
   END_RUNG
   // the same network as SCL:
   IF "UNO" THEN "DB124".Static_10 := FALSE; END_IF;
END_REGION

REGION Network 2
   RUNG wire#powerrail
      { S7_GenerateENO := "TRUE" } Move(in := 0, out1 => "DB121".Static_107)
   END_RUNG
   // the same network as SCL:
   "DB121".Static_107 := 0;
END_REGION

REGION Network 3
   RUNG wire#powerrail
      { S7_GenerateENO := "TRUE" } Move(in := 0, out1 => "DB121".Static_104)
   END_RUNG
   // the same network as SCL:
   "DB121".Static_104 := 0;
END_REGION

REGION Network 4
   RUNG wire#powerrail
      { S7_GenerateENO := "TRUE" } Move(in := -1, out1 => "DB121".Static_105)
   END_RUNG
   // the same network as SCL:
   "DB121".Static_105 := -1;
END_REGION

REGION Network 5
   RUNG wire#powerrail
      { S7_Templates := "SrcType := Int" } EQ_Contact(in1 := "DB124".Static_9, in2 := 0)
      wire#w1
      { S7_GenerateENO := "TRUE" } Move(in := 0, out1 => "DB121".Static_105)
   END_RUNG
   RUNG wire#w1
      S_Coil( "DB124".Static_10 )
   END_RUNG
   // the same network as SCL:
   IF "DB124".Static_9 = 0 THEN
       "DB121".Static_105 := 0;
       "DB124".Static_10 := TRUE;
   END_IF;
END_REGION

REGION Network 6
   IF NOT "DB124".Static_10 AND ("DB125".Static_1 = 1) AND "DB88".Static_12 THEN
       "DB121".Static_107 := "DB121".Static_107 + 1;
       "DB121".Static_104 := 1;
   END_IF;
END_REGION

REGION Network 7
   IF NOT "DB124".Static_10 AND ("DB121".Static_107 = "DB124".Static_9) THEN
       "DB121".Static_105 := 1;
       "DB124".Static_10 := TRUE;
   END_IF;
END_REGION

REGION Network 8
   IF NOT "DB124".Static_10 AND ("DB125".Static_2 = 1) AND "DB88".Static_13 THEN
       "DB121".Static_107 := "DB121".Static_107 + 1;
       "DB121".Static_104 := 1;
   END_IF;
END_REGION

REGION Network 9
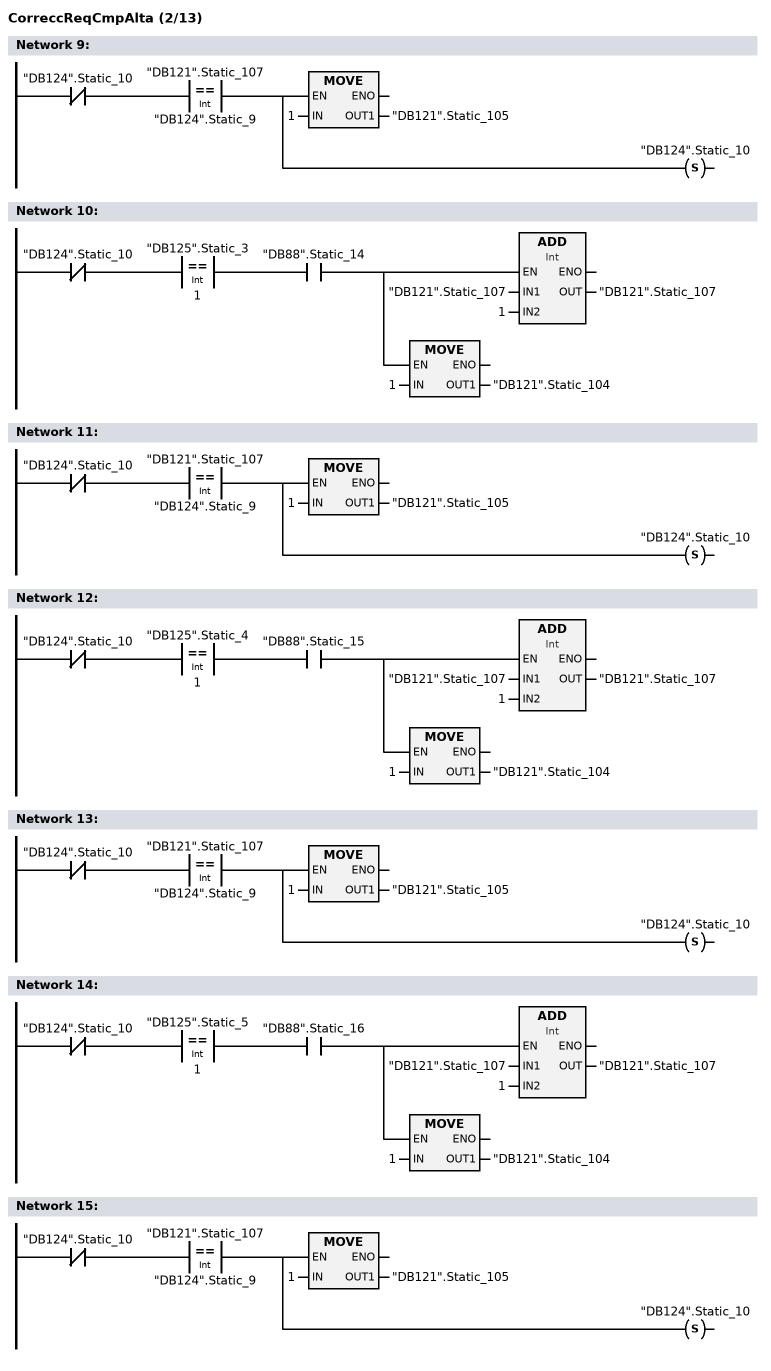
   IF NOT "DB124".Static_10 AND ("DB121".Static_107 = "DB124".Static_9) THEN
       "DB121".Static_105 := 1;
       "DB124".Static_10 := TRUE;
   END_IF;
END_REGION

REGION Network 10
   IF NOT "DB124".Static_10 AND ("DB125".Static_3 = 1) AND "DB88".Static_14 THEN
       "DB121".Static_107 := "DB121".Static_107 + 1;
       "DB121".Static_104 := 1;
   END_IF;
END_REGION

REGION Network 11
   IF NOT "DB124".Static_10 AND ("DB121".Static_107 = "DB124".Static_9) THEN
       "DB121".Static_105 := 1;
       "DB124".Static_10 := TRUE;
   END_IF;
END_REGION

REGION Network 12
   IF NOT "DB124".Static_10 AND ("DB125".Static_4 = 1) AND "DB88".Static_15 THEN
       "DB121".Static_107 := "DB121".Static_107 + 1;
       "DB121".Static_104 := 1;
   END_IF;
END_REGION

REGION Network 13
   IF NOT "DB124".Static_10 AND ("DB121".Static_107 = "DB124".Static_9) THEN
       "DB121".Static_105 := 1;
       "DB124".Static_10 := TRUE;
   END_IF;
END_REGION

REGION Network 14
   IF NOT "DB124".Static_10 AND ("DB125".Static_5 = 1) AND "DB88".Static_16 THEN
       "DB121".Static_107 := "DB121".Static_107 + 1;
       "DB121".Static_104 := 1;
   END_IF;
END_REGION

REGION Network 15
   IF NOT "DB124".Static_10 AND ("DB121".Static_107 = "DB124".Static_9) THEN
       "DB121".Static_105 := 1;
       "DB124".Static_10 := TRUE;
   END_IF;
END_REGION

REGION Network 16
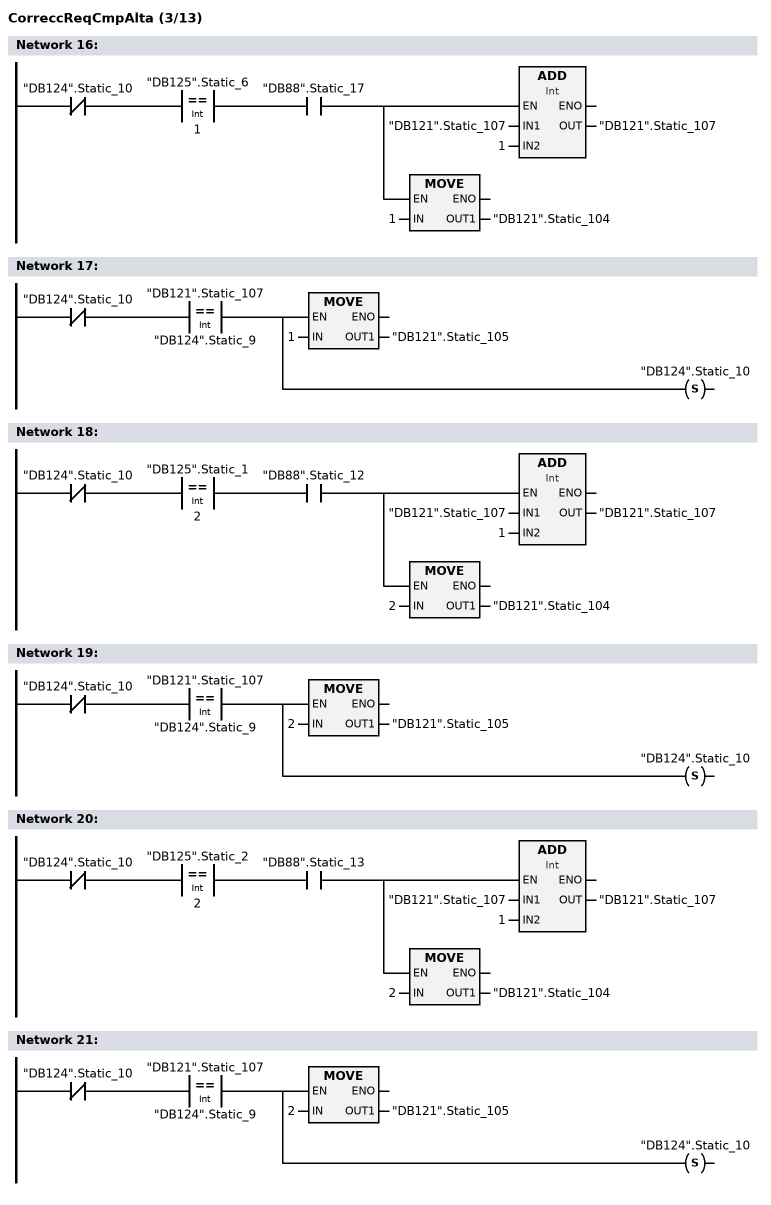
   IF NOT "DB124".Static_10 AND ("DB125".Static_6 = 1) AND "DB88".Static_17 THEN
       "DB121".Static_107 := "DB121".Static_107 + 1;
       "DB121".Static_104 := 1;
   END_IF;
END_REGION

REGION Network 17
   IF NOT "DB124".Static_10 AND ("DB121".Static_107 = "DB124".Static_9) THEN
       "DB121".Static_105 := 1;
       "DB124".Static_10 := TRUE;
   END_IF;
END_REGION

REGION Network 18
   IF NOT "DB124".Static_10 AND ("DB125".Static_1 = 2) AND "DB88".Static_12 THEN
       "DB121".Static_107 := "DB121".Static_107 + 1;
       "DB121".Static_104 := 2;
   END_IF;
END_REGION

REGION Network 19
   IF NOT "DB124".Static_10 AND ("DB121".Static_107 = "DB124".Static_9) THEN
       "DB121".Static_105 := 2;
       "DB124".Static_10 := TRUE;
   END_IF;
END_REGION

REGION Network 20
   IF NOT "DB124".Static_10 AND ("DB125".Static_2 = 2) AND "DB88".Static_13 THEN
       "DB121".Static_107 := "DB121".Static_107 + 1;
       "DB121".Static_104 := 2;
   END_IF;
END_REGION

REGION Network 21
   IF NOT "DB124".Static_10 AND ("DB121".Static_107 = "DB124".Static_9) THEN
       "DB121".Static_105 := 2;
       "DB124".Static_10 := TRUE;
   END_IF;
END_REGION

REGION Network 22
